FUNCTION_BLOCK "Vibrator B1"   // FB7, LAD
{ S7_Optimized_Access := 'TRUE' }
VERSION : 0.1
BEGIN

REGION Network 1
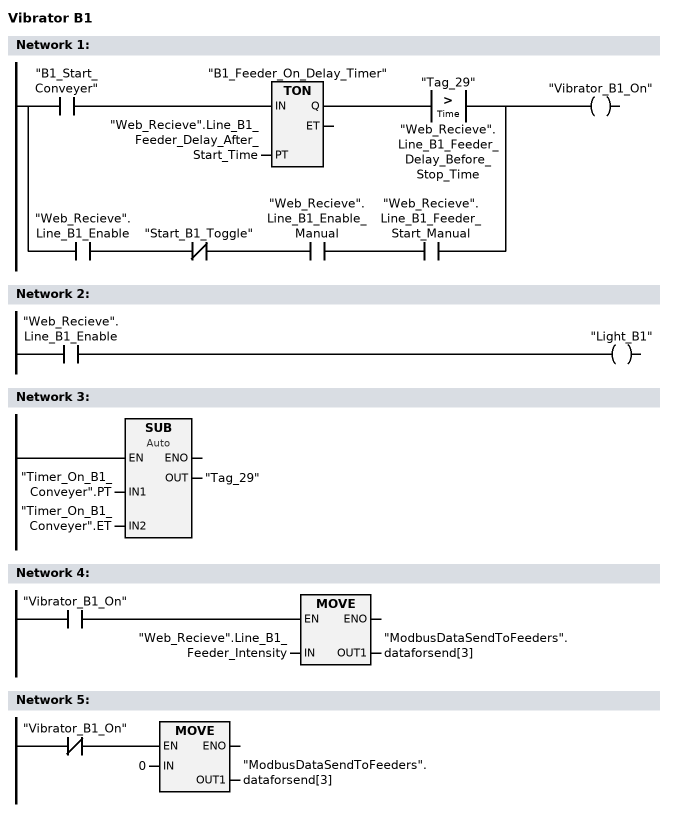
   "B1_Feeder_On_Delay_Timer".TON(IN := "B1_Start_Conveyer",
                           PT := "Web_Recieve".Line_B1_Feeder_Delay_After_Start_Time);
   "Vibrator_B1_On" := ("B1_Feeder_On_Delay_Timer".Q AND ("Tag_29" > "Web_Recieve".Line_B1_Feeder_Delay_Before_Stop_Time)) OR ("Web_Recieve".Line_B1_Enable AND NOT "Start_B1_Toggle" AND "Web_Recieve".Line_B1_Enable_Manual AND "Web_Recieve".Line_B1_Feeder_Start_Manual);
END_REGION

REGION Network 2
   RUNG wire#powerrail
      Contact( "Web_Recieve".Line_B1_Enable )
      Coil( "Light_B1" )
   END_RUNG
   // the same network as SCL:
   "Light_B1" := "Web_Recieve".Line_B1_Enable;
END_REGION

REGION Network 3
   RUNG wire#powerrail
      Sub(in1 := "Timer_On_B1_Conveyer".PT, in2 := "Timer_On_B1_Conveyer".ET, out => "Tag_29")
   END_RUNG
   // the same network as SCL:
   "Tag_29" := "Timer_On_B1_Conveyer".PT - "Timer_On_B1_Conveyer".ET;
END_REGION

REGION Network 4
   RUNG wire#powerrail
      Contact( "Vibrator_B1_On" )
      Move(in := "Web_Recieve".Line_B1_Feeder_Intensity, out1 => "ModbusDataSendToFeeders".dataforsend[3])
   END_RUNG
   // the same network as SCL:
   IF "Vibrator_B1_On" THEN
       "ModbusDataSendToFeeders".dataforsend[3] := "Web_Recieve".Line_B1_Feeder_Intensity;
   END_IF;
END_REGION

REGION Network 5
   RUNG wire#powerrail
      I_Contact( "Vibrator_B1_On" )
      Move(in := 0, out1 => "ModbusDataSendToFeeders".dataforsend[3])
   END_RUNG
   // the same network as SCL:
   IF NOT "Vibrator_B1_On" THEN "ModbusDataSendToFeeders".dataforsend[3] := 0; END_IF;
END_REGION
END_FUNCTION_BLOCK

FUNCTION_BLOCK "Vibrator B2"   // FB8, LAD
{ S7_Optimized_Access := 'TRUE' }
VERSION : 0.1
BEGIN

REGION Network 1
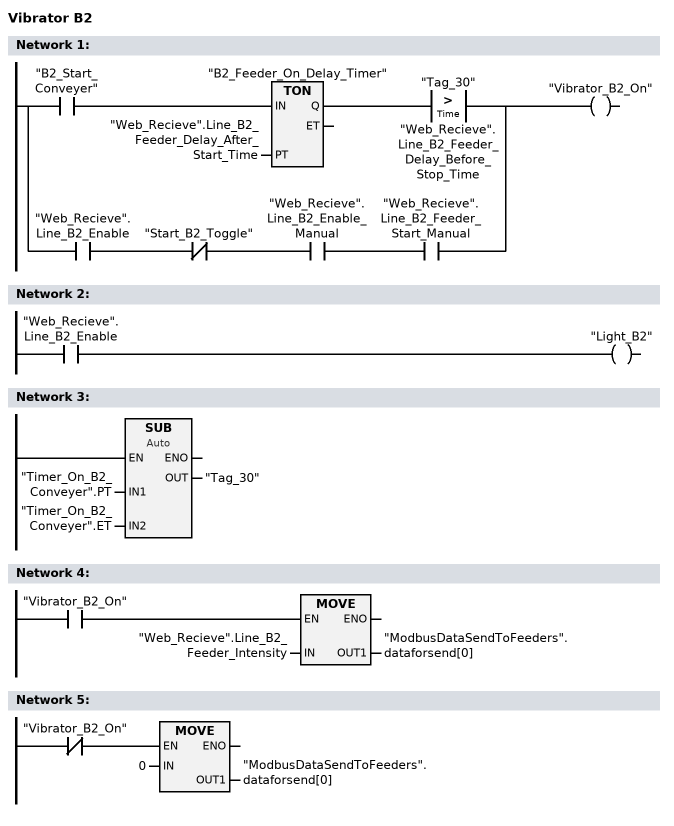
   "B2_Feeder_On_Delay_Timer".TON(IN := "B2_Start_Conveyer",
                           PT := "Web_Recieve".Line_B2_Feeder_Delay_After_Start_Time);
   "Vibrator_B2_On" := ("B2_Feeder_On_Delay_Timer".Q AND ("Tag_30" > "Web_Recieve".Line_B2_Feeder_Delay_Before_Stop_Time)) OR ("Web_Recieve".Line_B2_Enable AND NOT "Start_B2_Toggle" AND "Web_Recieve".Line_B2_Enable_Manual AND "Web_Recieve".Line_B2_Feeder_Start_Manual);
END_REGION

REGION Network 2
   RUNG wire#powerrail
      Contact( "Web_Recieve".Line_B2_Enable )
      Coil( "Light_B2" )
   END_RUNG
   // the same network as SCL:
   "Light_B2" := "Web_Recieve".Line_B2_Enable;
END_REGION

REGION Network 3
   RUNG wire#powerrail
      Sub(in1 := "Timer_On_B2_Conveyer".PT, in2 := "Timer_On_B2_Conveyer".ET, out => "Tag_30")
   END_RUNG
   // the same network as SCL:
   "Tag_30" := "Timer_On_B2_Conveyer".PT - "Timer_On_B2_Conveyer".ET;
END_REGION

REGION Network 4
   RUNG wire#powerrail
      Contact( "Vibrator_B2_On" )
      Move(in := "Web_Recieve".Line_B2_Feeder_Intensity, out1 => "ModbusDataSendToFeeders".dataforsend[0])
   END_RUNG
   // the same network as SCL:
   IF "Vibrator_B2_On" THEN
       "ModbusDataSendToFeeders".dataforsend[0] := "Web_Recieve".Line_B2_Feeder_Intensity;
   END_IF;
END_REGION

REGION Network 5
   RUNG wire#powerrail
      I_Contact( "Vibrator_B2_On" )
      Move(in := 0, out1 => "ModbusDataSendToFeeders".dataforsend[0])
   END_RUNG
   // the same network as SCL:
   IF NOT "Vibrator_B2_On" THEN "ModbusDataSendToFeeders".dataforsend[0] := 0; END_IF;
END_REGION
END_FUNCTION_BLOCK

FUNCTION_BLOCK "ConveyerA3_B3"   // FB9, LAD
{ S7_Optimized_Access := 'TRUE' }
VERSION : 0.1
BEGIN

REGION Network 1: Conveyor A3
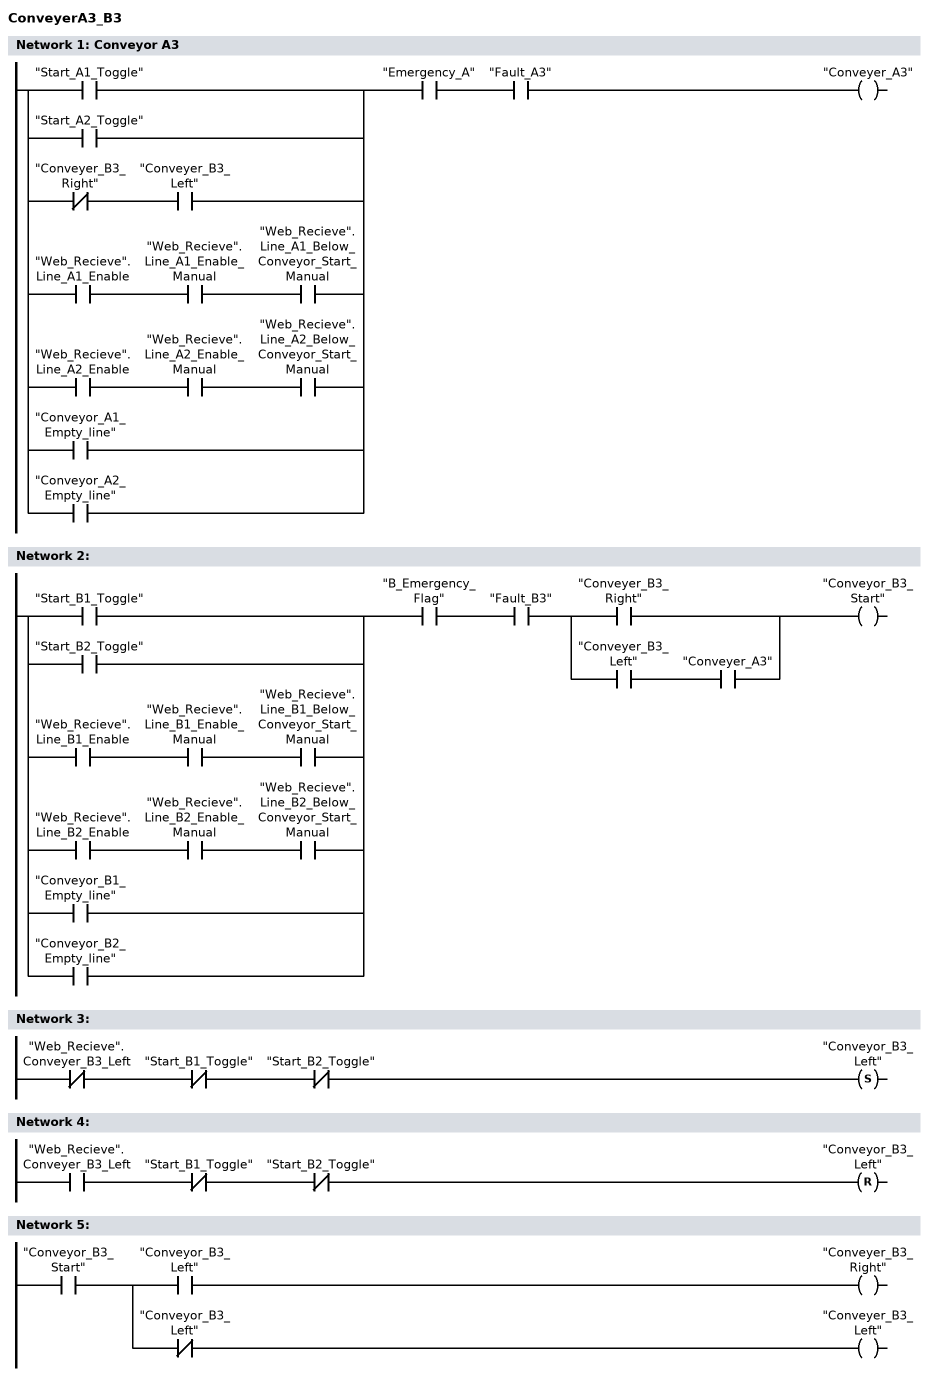
   RUNG wire#powerrail
      Contact( "Start_A1_Toggle" )
      wire#w1
      Contact( "Emergency_A" )
      Contact( "Fault_A3" )
      Coil( "Conveyer_A3" )
   END_RUNG
   RUNG wire#powerrail
      Contact( "Start_A2_Toggle" )
   END_RUNG wire#w1
   RUNG wire#powerrail
      I_Contact( "Conveyer_B3_Right" )
      Contact( "Conveyer_B3_Left" )
   END_RUNG wire#w1
   RUNG wire#powerrail
      Contact( "Web_Recieve".Line_A1_Enable )
      Contact( "Web_Recieve".Line_A1_Enable_Manual )
      Contact( "Web_Recieve".Line_A1_Below_Conveyor_Start_Manual )
   END_RUNG wire#w1
   RUNG wire#powerrail
      Contact( "Web_Recieve".Line_A2_Enable )
      Contact( "Web_Recieve".Line_A2_Enable_Manual )
      Contact( "Web_Recieve".Line_A2_Below_Conveyor_Start_Manual )
   END_RUNG wire#w1
   RUNG wire#powerrail
      Contact( "Conveyor_A1_Empty_line" )
   END_RUNG wire#w1
   RUNG wire#powerrail
      Contact( "Conveyor_A2_Empty_line" )
   END_RUNG wire#w1
   // the same network as SCL:
   "Conveyer_A3" := ("Start_A1_Toggle" OR "Start_A2_Toggle" OR (NOT "Conveyer_B3_Right" AND "Conveyer_B3_Left") OR ("Web_Recieve".Line_A1_Enable AND "Web_Recieve".Line_A1_Enable_Manual AND "Web_Recieve".Line_A1_Below_Conveyor_Start_Manual) OR ("Web_Recieve".Line_A2_Enable AND "Web_Recieve".Line_A2_Enable_Manual AND "Web_Recieve".Line_A2_Below_Conveyor_Start_Manual) OR "Conveyor_A1_Empty_line" OR "Conveyor_A2_Empty_line") AND "Emergency_A" AND "Fault_A3";
END_REGION

REGION Network 2
   RUNG wire#powerrail
      Contact( "Start_B1_Toggle" )
      wire#w1
      Contact( "B_Emergency_Flag" )
      Contact( "Fault_B3" )
      wire#w2
      Contact( "Conveyer_B3_Right" )
      wire#w3
      Coil( "Conveyor_B3_Start" )
   END_RUNG
   RUNG wire#powerrail
      Contact( "Start_B2_Toggle" )
   END_RUNG wire#w1
   RUNG wire#powerrail
      Contact( "Web_Recieve".Line_B1_Enable )
      Contact( "Web_Recieve".Line_B1_Enable_Manual )
      Contact( "Web_Recieve".Line_B1_Below_Conveyor_Start_Manual )
   END_RUNG wire#w1
   RUNG wire#powerrail
      Contact( "Web_Recieve".Line_B2_Enable )
      Contact( "Web_Recieve".Line_B2_Enable_Manual )
      Contact( "Web_Recieve".Line_B2_Below_Conveyor_Start_Manual )
   END_RUNG wire#w1
   RUNG wire#powerrail
      Contact( "Conveyor_B1_Empty_line" )
   END_RUNG wire#w1
   RUNG wire#powerrail
      Contact( "Conveyor_B2_Empty_line" )
   END_RUNG wire#w1
   RUNG wire#w2
      Contact( "Conveyer_B3_Left" )
      Contact( "Conveyer_A3" )
   END_RUNG wire#w3
   // the same network as SCL:
   "Conveyor_B3_Start" := ("Start_B1_Toggle" OR "Start_B2_Toggle" OR ("Web_Recieve".Line_B1_Enable AND "Web_Recieve".Line_B1_Enable_Manual AND "Web_Recieve".Line_B1_Below_Conveyor_Start_Manual) OR ("Web_Recieve".Line_B2_Enable AND "Web_Recieve".Line_B2_Enable_Manual AND "Web_Recieve".Line_B2_Below_Conveyor_Start_Manual) OR "Conveyor_B1_Empty_line" OR "Conveyor_B2_Empty_line") AND "B_Emergency_Flag" AND "Fault_B3" AND ("Conveyer_B3_Right" OR ("Conveyer_B3_Left" AND "Conveyer_A3"));
END_REGION

REGION Network 3
   RUNG wire#powerrail
      I_Contact( "Web_Recieve".Conveyer_B3_Left )
      I_Contact( "Start_B1_Toggle" )
      I_Contact( "Start_B2_Toggle" )
      S_Coil( "Conveyor_B3_Left" )
   END_RUNG
   // the same network as SCL:
   IF NOT "Web_Recieve".Conveyer_B3_Left AND NOT "Start_B1_Toggle" AND NOT "Start_B2_Toggle" THEN
       "Conveyor_B3_Left" := TRUE;
   END_IF;
END_REGION

REGION Network 4
   RUNG wire#powerrail
      Contact( "Web_Recieve".Conveyer_B3_Left )
      I_Contact( "Start_B1_Toggle" )
      I_Contact( "Start_B2_Toggle" )
      R_Coil( "Conveyor_B3_Left" )
   END_RUNG
   // the same network as SCL:
   IF "Web_Recieve".Conveyer_B3_Left AND NOT "Start_B1_Toggle" AND NOT "Start_B2_Toggle" THEN
       "Conveyor_B3_Left" := FALSE;
   END_IF;
END_REGION

REGION Network 5
   RUNG wire#powerrail
      Contact( "Conveyor_B3_Start" )
      wire#w1
      Contact( "Conveyor_B3_Left" )
      Coil( "Conveyer_B3_Right" )
   END_RUNG
   RUNG wire#w1
      I_Contact( "Conveyor_B3_Left" )
      Coil( "Conveyer_B3_Left" )
   END_RUNG
   // the same network as SCL:
   "Conveyer_B3_Right" := "Conveyor_B3_Start" AND "Conveyor_B3_Left";
   "Conveyer_B3_Left" := "Conveyor_B3_Start" AND NOT "Conveyor_B3_Left";
END_REGION
END_FUNCTION_BLOCK

FUNCTION_BLOCK "WebDataPrepaare"   // FB10, SCL
{ S7_Optimized_Access := 'TRUE' }
VERSION : 0.1
   VAR_TEMP
      WriteDBBusyTemp : Bool;
      writeresultValue : DInt;
   END_VAR
BEGIN
   "Web_Send".A_Emergency := NOT  "Emergency_A";
   "Web_Send".B_Emergency := NOT "Emergency_B";
   "Web_Send".A1_Conveyer := "Conveyer_A1";
   "Web_Send".A2_Conveyer := "Conveyer_A2";
   "Web_Send".B1_Conveyer := "Conveyer_B1";
   "Web_Send".B2_Conveyer := "Conveyer_B2";
   "Web_Send".A3_Conveyor := "Conveyer_A3";
   "Web_Send".B3_Left_Conveyer := NOT "Web_Recieve".Conveyer_B3_Left;
   "Web_Send".A1_Fault := NOT ("Fault_A1" AND "Fault_A3");
   "Web_Send".A2_Fault := NOT ("Fault_A2" AND "Fault_A3");
   "Web_Send".B1_Fault := NOT ("Fault_B1" AND "Fault_B3");
   "Web_Send".B2_Fault := NOT ("Fault_B2" AND "Fault_B3");
   "Web_Send".A1_Silo_Low := "Low_Silo_A1";
   "Web_Send".A2_Silo_Low := "Low_Silo_A2";
   "Web_Send".B1_Silo_Low := "Low_Silo_B1";
   "Web_Send".B2_Silo_Low := "Low_Silo_B2";
   "Web_Send".A1_Silo_High := "High_Silo_A1";
   "Web_Send".A2_Silo_High := "High_Silo_A2";
   "Web_Send".B1_Silo_High := "High_Silo_B1";
   "Web_Send".B2_Silo_High := "High_Silo_B2";
   "Web_Send".A1_Sample := "Pneumatic_A1";
   "Web_Send".A2_Sample := "Pneumatic_A2";
   "Web_Send".B1_Sample := "Pneumatic_B1";
   "Web_Send".B2_Sample := "Pneumatic_B2";
   "Web_Send".A1_Manual := "Web_Recieve".Line_A1_Enable_Manual;


   "Web_Send".A1_Running_Duration := "Web_Recieve".Line_A1_Conveyer_on_Time;
   "Web_Send".A1_Pause_Duration := "Web_Recieve".Line_A1_Conveyer_off_Time;
   "Web_Send".A1_Feeder_Vibration_Intensity := "Web_Recieve".Line_A1_Feeder_Intensity;
   "Web_Send".A1_Ruuning_Online := "Timer_Off_A1_Conveyer".PT - "Timer_Off_A1_Conveyer".ET;
   "Web_Send".A1_Pause_Online := "Timer_Off_A1_Conveyer".ET;
   "Web_Send".A1_Sample_Interval :="Web_Recieve".Line_A1_Sampling_Time;
   "Web_Send".A1_Sample_Duration := "Web_Recieve".Line_A1_Sampling_OpenTime;
   "Web_Send".A1_Sample_Online := "Timer_Before_On_Sample_A1".PT - "Timer_Before_On_Sample_A1".ET;
   "Web_Send".A1_Enable := "Web_Recieve".Line_A1_Enable;
   "Web_Send".A1_Start := "Start_A1_Toggle";
   "Web_Send".A1_Empty_Line_Time := "Web_Recieve".Line_A1_Empty_Line_Time;
   "Web_Send".A1_Feeder_Delay_After_Start_Time := "Web_Recieve".Line_A1_Feeder_Delay_After_Start_Time;
   "Web_Send".A1_Feeder_Delay_Before_Stop_Time := "Web_Recieve".Line_A1_Feeder_Delay_Before_Stop_Time;
   "Web_Send".A1_Duration_Big_Silo_Stop_Time := "Web_Recieve".Line_A1_Big_Silo_Delay_Start;

   "Web_Send".A2_Running_Duration := "Web_Recieve".Line_A2_Conveyer_on_Time;
   "Web_Send".A2_Pause_Duration := "Web_Recieve".Line_A2_Conveyer_off_Time;
   "Web_Send".A2_Feeder_Vibration_Intensity := "Web_Recieve".Line_A2_Feeder_Intensity;
   "Web_Send".A2_Ruuning_Online := "Timer_Off_A2_Conveyer".PT - "Timer_Off_A2_Conveyer".ET;
   "Web_Send".A2_Pause_Online := "Timer_Off_A2_Conveyer".ET;
   "Web_Send".A2_Sample_Interval := "Web_Recieve".Line_A2_Sampling_Time;
   "Web_Send".A2_Sample_Duration := "Web_Recieve".Line_A2_Sampling_OpenTime;
   "Web_Send".A2_Sample_Online := "Timer_Before_On_Sample_A2".PT - "Timer_Before_On_Sample_A2".ET;
   "Web_Send".A2_Enable := "Web_Recieve".Line_A2_Enable;
   "Web_Send".A2_Start := "Start_A2_Toggle";
   "Web_Send".A2_Empty_Line_Time := "Web_Recieve".Line_A2_Empty_Line_Time;
   "Web_Send".A2_Feeder_Delay_After_Start_Time := "Web_Recieve".Line_A2_Feeder_Delay_After_Start_Time;
   "Web_Send".A2_Feeder_Delay_Before_Stop_Time := "Web_Recieve".Line_A2_Feeder_Delay_Before_Stop_Time;
   "Web_Send".A2_Duration_Big_Silo_Stop_Time := "Web_Recieve".Line_A2_Big_Silo_Delay_Start;


   "Web_Send".B1_Running_Duration := "Web_Recieve".Line_B1_Conveyer_on_Time;
   "Web_Send".B1_Pause_Duration := "Web_Recieve".Line_B1_Conveyer_off_Time;
   "Web_Send".B1_Feeder_Vibration_Intensity := "Web_Recieve".Line_B1_Feeder_Intensity;
   "Web_Send".B1_Ruuning_Online := "Timer_On_B1_Conveyer".ET;
   "Web_Send".B1_Pause_Online := "Timer_Off_B1_Conveyer".ET;
   "Web_Send".B1_Sample_Interval := "Web_Recieve".Line_B1_Sampling_Time;
   "Web_Send".B1_Sample_Duration := "Web_Recieve".Line_B1_Sampling_OpenTime;
   "Web_Send".B1_Sample_Online := "Timer_Before_On_Sample_B1".ET - "Timer_Before_On_Sample_B1".ET;
   "Web_Send".B1_Enable := "Web_Recieve".Line_B1_Enable;
   "Web_Send".B1_Start := "Start_B1_Toggle";
   "Web_Send".B1_Empty_Line_Time := "Web_Recieve".Line_B1_Empty_Line_Time;
   "Web_Send".B1_Feeder_Delay_After_Start_Time := "Web_Recieve".Line_B1_Feeder_Delay_After_Start_Time;
   "Web_Send".B1_Feeder_Delay_Before_Stop_Time := "Web_Recieve".Line_B1_Feeder_Delay_Before_Stop_Time;
   "Web_Send".B1_Duration_Big_Silo_Stop_Time := "Web_Recieve".Line_B1_Big_Silo_Delay_Start;


   "Web_Send".B2_Running_Duration := "Web_Recieve".Line_B2_Conveyer_on_Time;
   "Web_Send".B2_Pause_Duration := "Web_Recieve".Line_B2_Conveyer_off_Time;
   "Web_Send".B2_Feeder_Vibration_Intensity := "Web_Recieve".Line_B2_Feeder_Intensity;
   "Web_Send".B2_Ruuning_Online := "Timer_On_B2_Conveyer".ET;
   "Web_Send".B2_Pause_Online := "Timer_Off_B2_Conveyer".ET;
   "Web_Send".B2_Sample_Interval := "Web_Recieve".Line_B2_Sampling_Time;
   "Web_Send".B2_Sample_Duration := "Web_Recieve".Line_B2_Sampling_OpenTime;
   "Web_Send".B2_Sample_Online := "Timer_Before_On_Sample_B2".ET - "Timer_Before_On_Sample_B2".ET;
   "Web_Send".B2_Enable := "Web_Recieve".Line_B2_Enable;
   "Web_Send".B2_Start := "Start_B2_Toggle";
   "Web_Send".B2_Empty_Line_Time := "Web_Recieve".Line_B2_Empty_Line_Time;
   "Web_Send".B2_Feeder_Delay_After_Start_Time := "Web_Recieve".Line_B2_Feeder_Delay_After_Start_Time;
   "Web_Send".B2_Feeder_Delay_Before_Stop_Time := "Web_Recieve".Line_B2_Feeder_Delay_Before_Stop_Time;
   "Web_Send".B2_Duration_Big_Silo_Stop_Time := "Web_Recieve".Line_B2_Big_Silo_Delay_Start;
END_FUNCTION_BLOCK

FUNCTION_BLOCK "Sample"   // FB11, LAD
{ S7_Optimized_Access := 'TRUE' }
VERSION : 0.1
   VAR_TEMP   // added for the SCL form of the ladder/FBD networks
      _w1 : Bool;
   END_VAR
BEGIN

REGION Network 1: A1 Before Sample
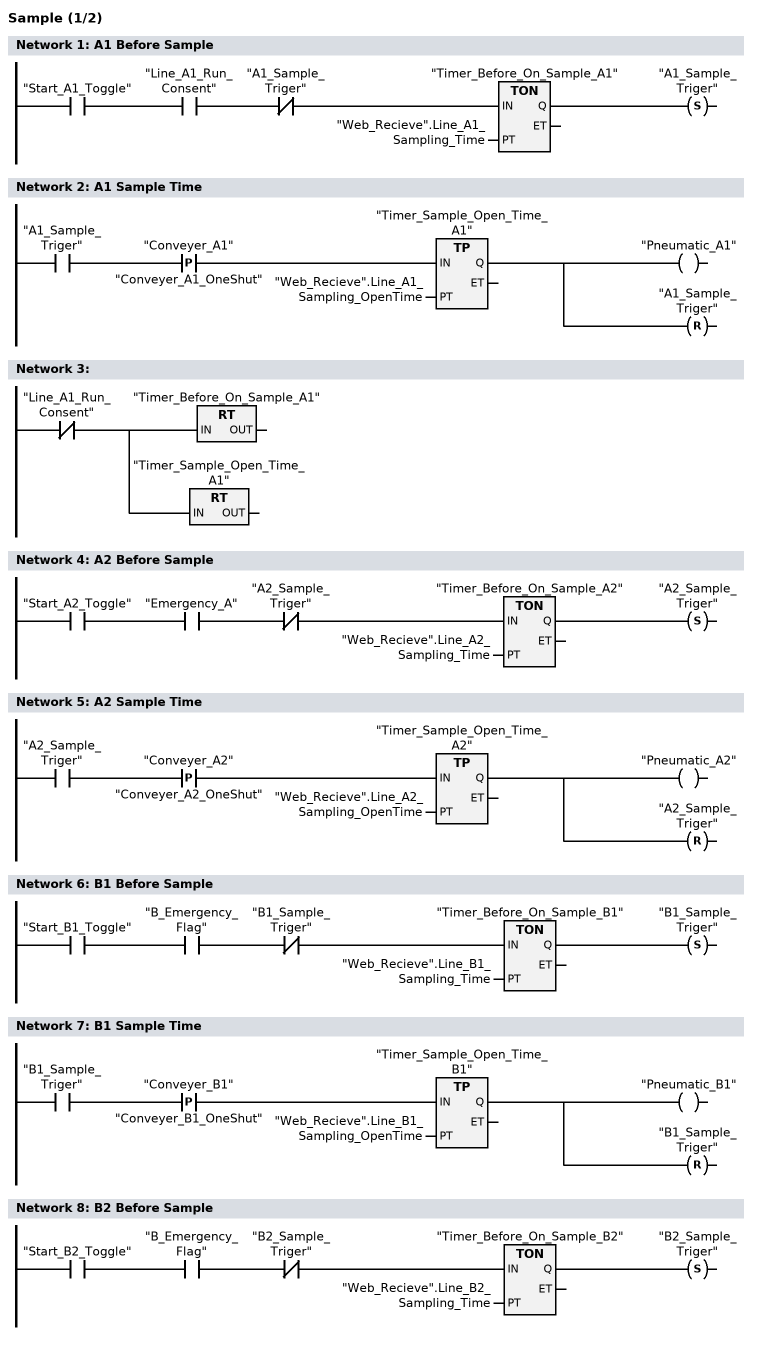
   "Timer_Before_On_Sample_A1".TON(IN := "Start_A1_Toggle" AND "Line_A1_Run_Consent" AND NOT "A1_Sample_Triger",
                           PT := "Web_Recieve".Line_A1_Sampling_Time);
   IF "Timer_Before_On_Sample_A1".Q THEN "A1_Sample_Triger" := TRUE; END_IF;
END_REGION

REGION Network 2: A1 Sample Time
   #_w1 := "A1_Sample_Triger" AND "Conveyer_A1" AND NOT "Conveyer_A1_OneShut";   // rising edge of "Conveyer_A1"
   "Conveyer_A1_OneShut" := "Conveyer_A1";
   "Timer_Sample_Open_Time_A1".TP(IN := #_w1, PT := "Web_Recieve".Line_A1_Sampling_OpenTime);
   "Pneumatic_A1" := "Timer_Sample_Open_Time_A1".Q;
   IF "Timer_Sample_Open_Time_A1".Q THEN "A1_Sample_Triger" := FALSE; END_IF;
END_REGION

REGION Network 3
   RUNG wire#powerrail
      I_Contact( "Line_A1_Run_Consent" )
      wire#w1
      RT_Coil( "Timer_Before_On_Sample_A1" )
   END_RUNG
   RUNG wire#w1
      RT_Coil( "Timer_Sample_Open_Time_A1" )
   END_RUNG
   // the same network as SCL:
   #_w1 := NOT "Line_A1_Run_Consent";
   IF #_w1 THEN
       RESET_TIMER("Timer_Before_On_Sample_A1");
       RESET_TIMER("Timer_Sample_Open_Time_A1");
   END_IF;
END_REGION

REGION Network 4: A2 Before Sample
   "Timer_Before_On_Sample_A2".TON(IN := "Start_A2_Toggle" AND "Emergency_A" AND NOT "A2_Sample_Triger",
                           PT := "Web_Recieve".Line_A2_Sampling_Time);
   IF "Timer_Before_On_Sample_A2".Q THEN "A2_Sample_Triger" := TRUE; END_IF;
END_REGION

REGION Network 5: A2 Sample Time
   #_w1 := "A2_Sample_Triger" AND "Conveyer_A2" AND NOT "Conveyer_A2_OneShut";   // rising edge of "Conveyer_A2"
   "Conveyer_A2_OneShut" := "Conveyer_A2";
   "Timer_Sample_Open_Time_A2".TP(IN := #_w1, PT := "Web_Recieve".Line_A2_Sampling_OpenTime);
   "Pneumatic_A2" := "Timer_Sample_Open_Time_A2".Q;
   IF "Timer_Sample_Open_Time_A2".Q THEN "A2_Sample_Triger" := FALSE; END_IF;
END_REGION

REGION Network 6: B1 Before Sample
   "Timer_Before_On_Sample_B1".TON(IN := "Start_B1_Toggle" AND "B_Emergency_Flag" AND NOT "B1_Sample_Triger",
                           PT := "Web_Recieve".Line_B1_Sampling_Time);
   IF "Timer_Before_On_Sample_B1".Q THEN "B1_Sample_Triger" := TRUE; END_IF;
END_REGION

REGION Network 7: B1 Sample Time
   #_w1 := "B1_Sample_Triger" AND "Conveyer_B1" AND NOT "Conveyer_B1_OneShut";   // rising edge of "Conveyer_B1"
   "Conveyer_B1_OneShut" := "Conveyer_B1";
   "Timer_Sample_Open_Time_B1".TP(IN := #_w1, PT := "Web_Recieve".Line_B1_Sampling_OpenTime);
   "Pneumatic_B1" := "Timer_Sample_Open_Time_B1".Q;
   IF "Timer_Sample_Open_Time_B1".Q THEN "B1_Sample_Triger" := FALSE; END_IF;
END_REGION

REGION Network 8: B2 Before Sample
   "Timer_Before_On_Sample_B2".TON(IN := "Start_B2_Toggle" AND "B_Emergency_Flag" AND NOT "B2_Sample_Triger",
                           PT := "Web_Recieve".Line_B2_Sampling_Time);
   IF "Timer_Before_On_Sample_B2".Q THEN "B2_Sample_Triger" := TRUE; END_IF;
END_REGION

REGION Network 9: B2 Sample Time
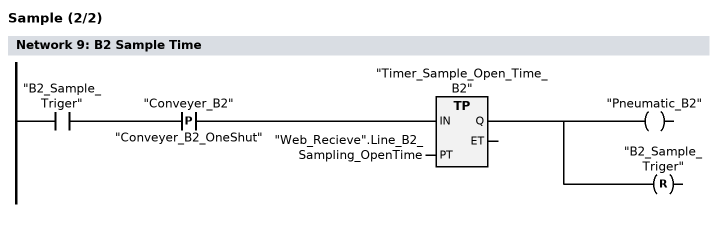
   #_w1 := "B2_Sample_Triger" AND "Conveyer_B2" AND NOT "Conveyer_B2_OneShut";   // rising edge of "Conveyer_B2"
   "Conveyer_B2_OneShut" := "Conveyer_B2";
   "Timer_Sample_Open_Time_B2".TP(IN := #_w1, PT := "Web_Recieve".Line_B2_Sampling_OpenTime);
   "Pneumatic_B2" := "Timer_Sample_Open_Time_B2".Q;
   IF "Timer_Sample_Open_Time_B2".Q THEN "B2_Sample_Triger" := FALSE; END_IF;
END_REGION
END_FUNCTION_BLOCK

FUNCTION_BLOCK "Silo_Big_A-B"   // FB12, LAD
{ S7_Optimized_Access := 'TRUE' }
VERSION : 0.1
BEGIN

REGION Network 1
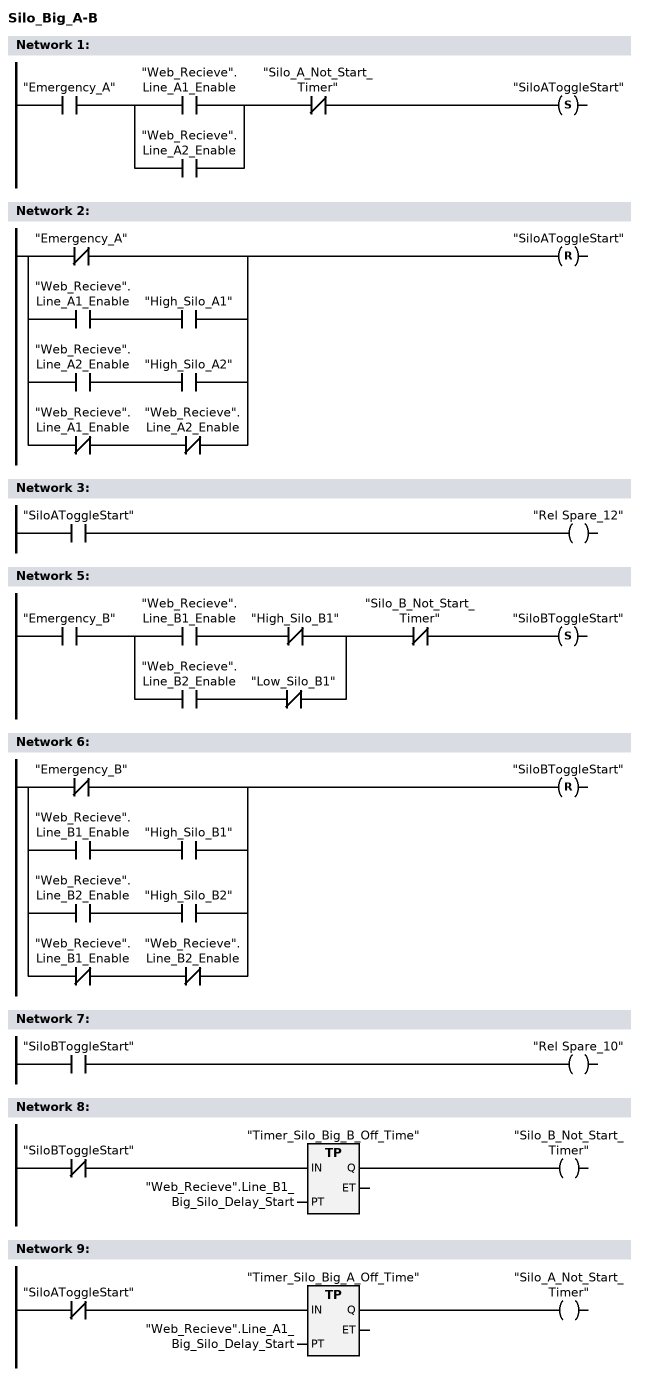
   RUNG wire#powerrail
      Contact( "Emergency_A" )
      wire#w1
      Contact( "Web_Recieve".Line_A1_Enable )
      wire#w2
      I_Contact( "Silo_A_Not_Start_Timer" )
      S_Coil( "SiloAToggleStart" )
   END_RUNG
   RUNG wire#w1
      Contact( "Web_Recieve".Line_A2_Enable )
   END_RUNG wire#w2
   // the same network as SCL:
   IF "Emergency_A" AND ("Web_Recieve".Line_A1_Enable OR "Web_Recieve".Line_A2_Enable) AND NOT "Silo_A_Not_Start_Timer" THEN
       "SiloAToggleStart" := TRUE;
   END_IF;
END_REGION

REGION Network 2
   RUNG wire#powerrail
      I_Contact( "Emergency_A" )
      wire#w1
      R_Coil( "SiloAToggleStart" )
   END_RUNG
   RUNG wire#powerrail
      Contact( "Web_Recieve".Line_A1_Enable )
      Contact( "High_Silo_A1" )
   END_RUNG wire#w1
   RUNG wire#powerrail
      Contact( "Web_Recieve".Line_A2_Enable )
      Contact( "High_Silo_A2" )
   END_RUNG wire#w1
   RUNG wire#powerrail
      I_Contact( "Web_Recieve".Line_A1_Enable )
      I_Contact( "Web_Recieve".Line_A2_Enable )
   END_RUNG wire#w1
   // the same network as SCL:
   IF NOT "Emergency_A" OR ("Web_Recieve".Line_A1_Enable AND "High_Silo_A1") OR ("Web_Recieve".Line_A2_Enable AND "High_Silo_A2") OR (NOT "Web_Recieve".Line_A1_Enable AND NOT "Web_Recieve".Line_A2_Enable) THEN
       "SiloAToggleStart" := FALSE;
   END_IF;
END_REGION

REGION Network 3
   RUNG wire#powerrail
      Contact( "SiloAToggleStart" )
      Coil( "Rel Spare_12" )
   END_RUNG
   // the same network as SCL:
   "Rel Spare_12" := "SiloAToggleStart";
END_REGION

REGION Network 5
   RUNG wire#powerrail
      Contact( "Emergency_B" )
      wire#w1
      Contact( "Web_Recieve".Line_B1_Enable )
      I_Contact( "High_Silo_B1" )
      wire#w2
      I_Contact( "Silo_B_Not_Start_Timer" )
      S_Coil( "SiloBToggleStart" )
   END_RUNG
   RUNG wire#w1
      Contact( "Web_Recieve".Line_B2_Enable )
      I_Contact( "Low_Silo_B1" )
   END_RUNG wire#w2
   // the same network as SCL:
   IF "Emergency_B" AND (("Web_Recieve".Line_B1_Enable AND NOT "High_Silo_B1") OR ("Web_Recieve".Line_B2_Enable AND NOT "Low_Silo_B1")) AND NOT "Silo_B_Not_Start_Timer" THEN
       "SiloBToggleStart" := TRUE;
   END_IF;
END_REGION

REGION Network 6
   RUNG wire#powerrail
      I_Contact( "Emergency_B" )
      wire#w1
      R_Coil( "SiloBToggleStart" )
   END_RUNG
   RUNG wire#powerrail
      Contact( "Web_Recieve".Line_B1_Enable )
      Contact( "High_Silo_B1" )
   END_RUNG wire#w1
   RUNG wire#powerrail
      Contact( "Web_Recieve".Line_B2_Enable )
      Contact( "High_Silo_B2" )
   END_RUNG wire#w1
   RUNG wire#powerrail
      I_Contact( "Web_Recieve".Line_B1_Enable )
      I_Contact( "Web_Recieve".Line_B2_Enable )
   END_RUNG wire#w1
   // the same network as SCL:
   IF NOT "Emergency_B" OR ("Web_Recieve".Line_B1_Enable AND "High_Silo_B1") OR ("Web_Recieve".Line_B2_Enable AND "High_Silo_B2") OR (NOT "Web_Recieve".Line_B1_Enable AND NOT "Web_Recieve".Line_B2_Enable) THEN
       "SiloBToggleStart" := FALSE;
   END_IF;
END_REGION

REGION Network 7
   RUNG wire#powerrail
      Contact( "SiloBToggleStart" )
      Coil( "Rel Spare_10" )
   END_RUNG
   // the same network as SCL:
   "Rel Spare_10" := "SiloBToggleStart";
END_REGION

REGION Network 8
   "Timer_Silo_Big_B_Off_Time".TP(IN := NOT "SiloBToggleStart",
                           PT := "Web_Recieve".Line_B1_Big_Silo_Delay_Start);
   "Silo_B_Not_Start_Timer" := "Timer_Silo_Big_B_Off_Time".Q;
END_REGION

REGION Network 9
   "Timer_Silo_Big_A_Off_Time".TP(IN := NOT "SiloAToggleStart",
                           PT := "Web_Recieve".Line_A1_Big_Silo_Delay_Start);
   "Silo_A_Not_Start_Timer" := "Timer_Silo_Big_A_Off_Time".Q;
END_REGION
END_FUNCTION_BLOCK

FUNCTION_BLOCK "Empty Line A1 A2"   // FB13, LAD
{ S7_Optimized_Access := 'TRUE' }
VERSION : 0.1
   VAR_TEMP   // added for the SCL form of the ladder/FBD networks
      _w1 : Bool;
   END_VAR
BEGIN

REGION Network 1: Empty Line A1